(* Logix 5000 project; controller _GigaDiscovery vendor 1 type 14 code 244 rev 35.11; software revision 35.03; part 8 of 23 *)
(* tags used below, declared in another part *)
   ArmInductanceGondola : REAL;
   ArmResistanceGondola : REAL;
   First_Push_Angle : REAL;   // WEIGHT
   Gondola_Start_Delay : TIMER;
   Gondola_Stop : BOOL;
   Max_Torque_for_Angle_Correction : REAL;
   Min_error_to_Start_Decreasing_Torque : REAL;
   Os : DINT;
   Os_to_CCW : BOOL;
   Os_to_CW : BOOL;
   Pylon_Sequencer : Sequencer;
   SpeedRegKi : REAL;
   SpeedRegKp : REAL;
   Timer : TIMER[10];
   Angle_at_Full_Load : REAL;
   Angle_at_min_Load : REAL;
   AngleContrl : REAL;
   Auto_Cycle_Step : DINT;
   Braking_Torque_Lim : REAL;
   CurrentLimit : DINT;
   Direction : BOOL;   // 1 = Spinta CW 0 = Spinta CCW
   Enable_to_Start : UDT_CROUT;   // Abilitazione allo start QC8011E QC8013E
   Encoder_Resetted : BOOL;
   First_Push_Set_Torque_to_Zero : BOOL;
   Girella_Field_Actuate_During_Inactivity : BOOL;
   Gondola_Axe : Axe;
   Gondola_Decc_timer_Start : BOOL;
   Gondola_Immediatly_Stop : BOOL;
   Gondola_Out_Ref : INT;
   Gondola_Speed_Ref_ABS : REAL;
   Gondola_Speed_Reference : DINT;
   Gondola_Stop_CW : BOOL;   // Gondola Sto Direction 0 > CCW 1 > CW
   Gondola_Stop_Step : DINT;
   HMI_Gondola_Start_Delay : DINT;
   HMI_Overspeed_Test_Pb : BOOL;
   HMI_Reset_Encoder_Position : BOOL;
   I_Gondola_Home_Position_Sensor_1 : UDT_DCM;   // Home Sensor Speed Check -B40002I
   I_Pylon_Home_Ch1 : UDT_DCM;   // Home position Pylon Ch1 -B26002I
   I_Pylon_Home_Ch2 : UDT_DCM;   // Home position Pylon Ch2 -B26007I
   I_Zero_Set_Sensor : BOOL;   // Zero Set Sensor -B11201A
   Increase_Torque_Limit_Mem : BOOL;
   K_Brake : REAL;
   K_Speed_Factor : REAL;
   Max_Empty_Torque : REAL;   // 75
   Max_Full_Torque : REAL;   // 85
   MAX_HMI_Speed_Value : DINT;
   Max_Reference_Output : DINT;
   Max_Speed_Reference : DINT;
   Min_Speed_Reference : DINT;
   Min_Torque_to_Maintain_Height_Full_Load : REAL;
   Min_Torque_to_Maintain_Height_min_Load : REAL;
   No_Sfty : Std_to_Sfty;
   Os_to_CW_CCW : BOOL;
   Oscillation_Error : REAL;
   Pylon_Axe : Axe;
   Pylon_Field_Actuate_During_Inactivity : BOOL;
   Pylon_Filtered_Speed : REAL;
   Pylon_Reference : DINT;
   Ratio_HMI_Speed_Ref : REAL;
   Reference_Out_Conversion_Pylon : REAL;
   Reset_Pulse : BOOL;
   RPM_Max_Motor_Speed_Pylon : DINT;
   Start_Stop_Cycle : Sequencer;
   Stop_Request : BOOL;
   Timers : TIMER[32];
   To_Sfty : Std_to_Sfty;
   Torque_Cmd_from_Cycle : REAL;
   TorqueNeg_Angle_Control : REAL;
   TorquePos_Angle_Control : REAL;
   Work_Auto_Cycle : Auto_Cycle;
(* Pylon, continued *)

ROUTINE _02_Ctrl_Mode   (* ladder *)
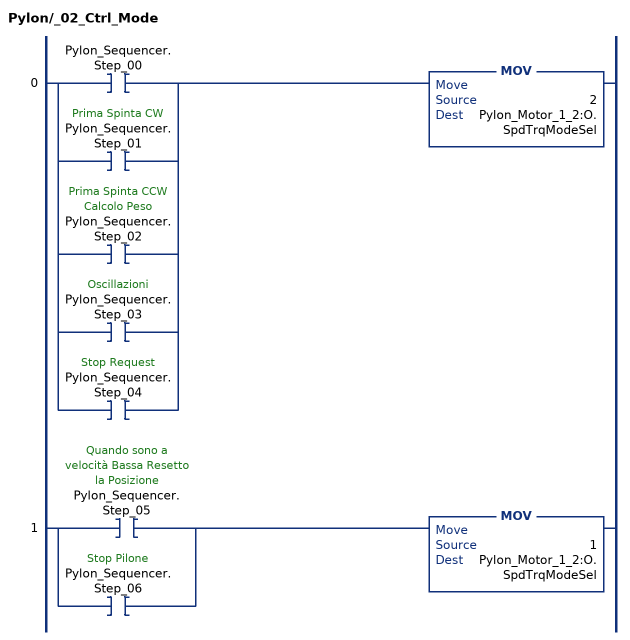
   0: [XIC(Pylon_Sequencer.Step_00) ,XIC(Pylon_Sequencer.Step_01) ,XIC(Pylon_Sequencer.Step_02) ,XIC(Pylon_Sequencer.Step_03) ,XIC(Pylon_Sequencer.Step_04) ]MOV(2,Pylon_Motor_1_2:O.SpdTrqModeSel);
   1: [XIC(Pylon_Sequencer.Step_05) ,XIC(Pylon_Sequencer.Step_06) ]MOV(1,Pylon_Motor_1_2:O.SpdTrqModeSel);
END_ROUTINE

ROUTINE _03_Speed_Ref   (* ladder *)
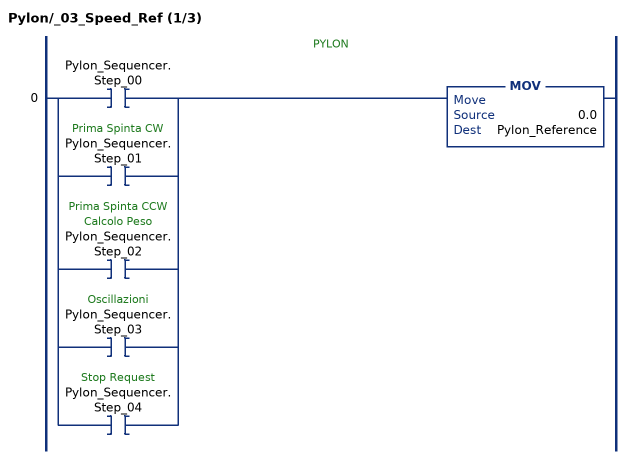
   // PYLON
   0: [XIC(Pylon_Sequencer.Step_00) ,XIC(Pylon_Sequencer.Step_01) ,XIC(Pylon_Sequencer.Step_02) ,XIC(Pylon_Sequencer.Step_03) ,XIC(Pylon_Sequencer.Step_04) ]MOV(0.0,Pylon_Reference);
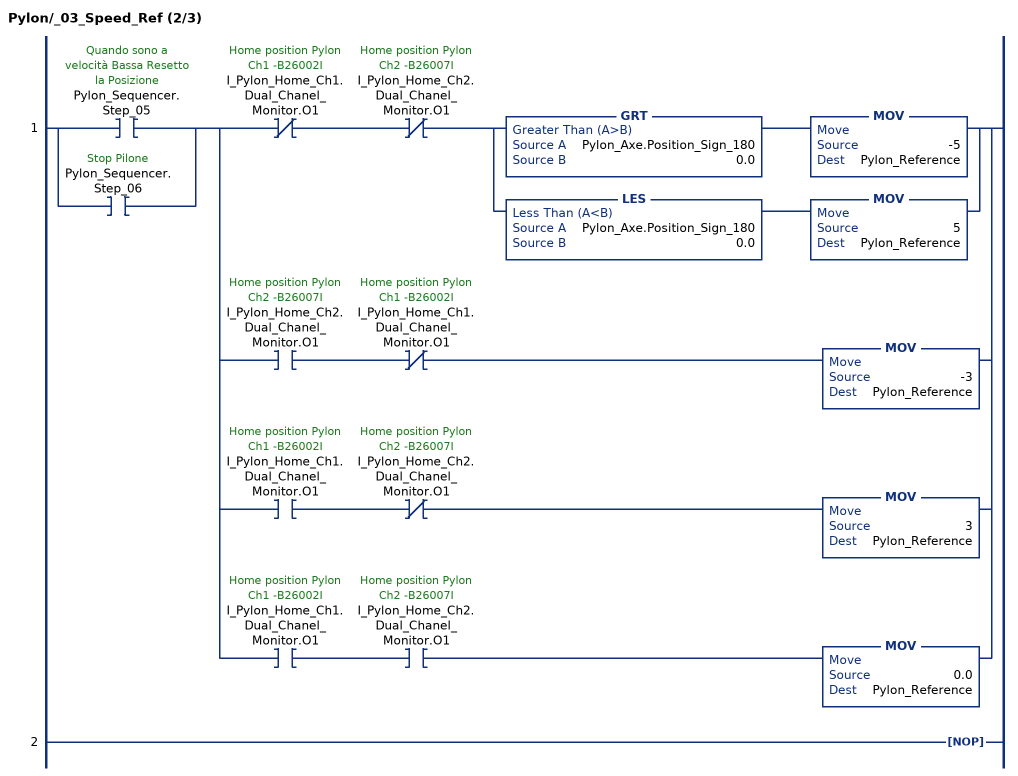
   1: [XIC(Pylon_Sequencer.Step_05) ,XIC(Pylon_Sequencer.Step_06) ][XIO(I_Pylon_Home_Ch1.Dual_Chanel_Monitor.O1) XIO(I_Pylon_Home_Ch2.Dual_Chanel_Monitor.O1) [GRT(Pylon_Axe.Position_Sign_180,0.0) MOV(-5,Pylon_Reference) ,LES(Pylon_Axe.Position_Sign_180,0.0) MOV(5,Pylon_Reference) ] ,[XIC(I_Pylon_Home_Ch2.Dual_Chanel_Monitor.O1) XIO(I_Pylon_Home_Ch1.Dual_Chanel_Monitor.O1) MOV(-3,Pylon_Reference) ,XIC(I_Pylon_Home_Ch1.Dual_Chanel_Monitor.O1) XIO(I_Pylon_Home_Ch2.Dual_Chanel_Monitor.O1) MOV(3,Pylon_Reference) ,XIC(I_Pylon_Home_Ch1.Dual_Chanel_Monitor.O1) XIC(I_Pylon_Home_Ch2.Dual_Chanel_Monitor.O1) MOV(0.0,Pylon_Reference) ] ];
   2: NOP();
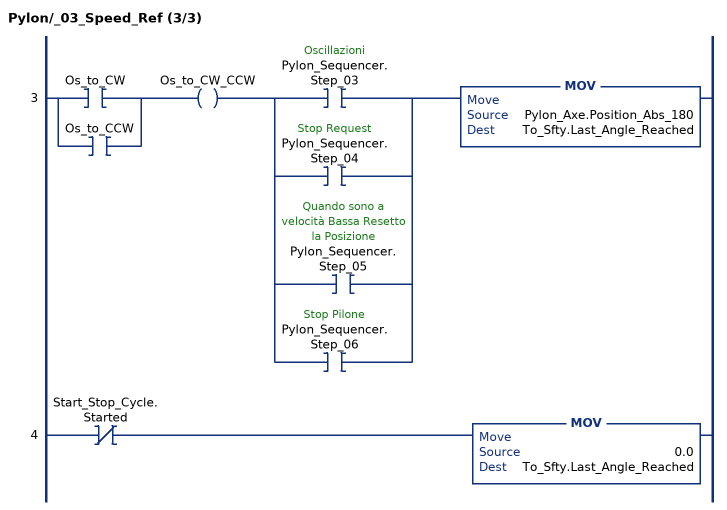
   3: [XIC(Os_to_CW) ,XIC(Os_to_CCW) ]OTE(Os_to_CW_CCW)[XIC(Pylon_Sequencer.Step_03) ,XIC(Pylon_Sequencer.Step_04) ,XIC(Pylon_Sequencer.Step_05) ,XIC(Pylon_Sequencer.Step_06) ]MOV(Pylon_Axe.Position_Abs_180,To_Sfty.Last_Angle_Reached);
   4: XIO(Start_Stop_Cycle.Started)MOV(0.0,To_Sfty.Last_Angle_Reached);
END_ROUTINE

ROUTINE _04_Torque_Lim   (* ladder *)
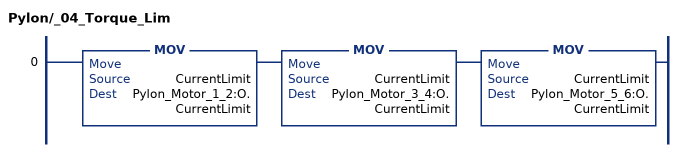
   0: MOV(CurrentLimit,Pylon_Motor_1_2:O.CurrentLimit)MOV(CurrentLimit,Pylon_Motor_3_4:O.CurrentLimit)MOV(CurrentLimit,Pylon_Motor_5_6:O.CurrentLimit);
END_ROUTINE

ROUTINE _05_Oscillation   (* ladder *)
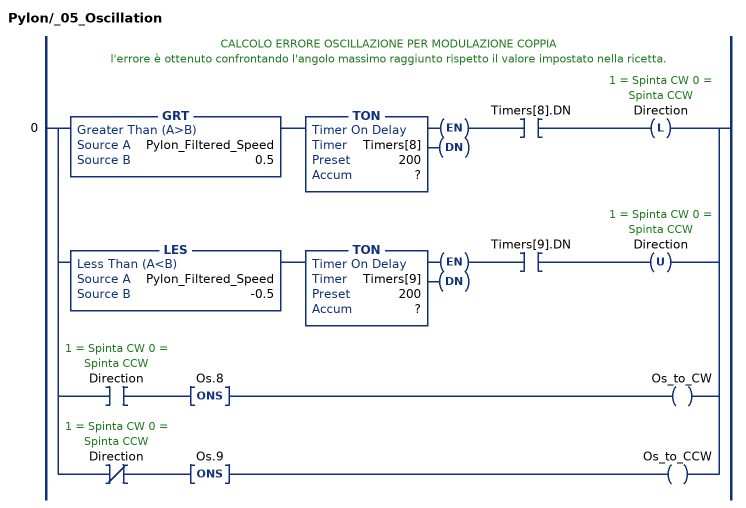
   // CALCOLO ERRORE OSCILLAZIONE PER MODULAZIONE COPPIA
   // l'errore è ottenuto confrontando l'angolo massimo raggiunto rispetto il valore impostato nella ricetta.
   0: [GRT(Pylon_Filtered_Speed,0.5) TON(Timers[8],?,?) XIC(Timers[8].DN) OTL(Direction) ,LES(Pylon_Filtered_Speed,-0.5) TON(Timers[9],?,?) XIC(Timers[9].DN) OTU(Direction) ,XIC(Direction) ONS(Os.8) OTE(Os_to_CW) ,XIO(Direction) ONS(Os.9) OTE(Os_to_CCW) ];
END_ROUTINE

ROUTINE _06_Scale_Angle   (* function block diagram *)
   SHEET 1
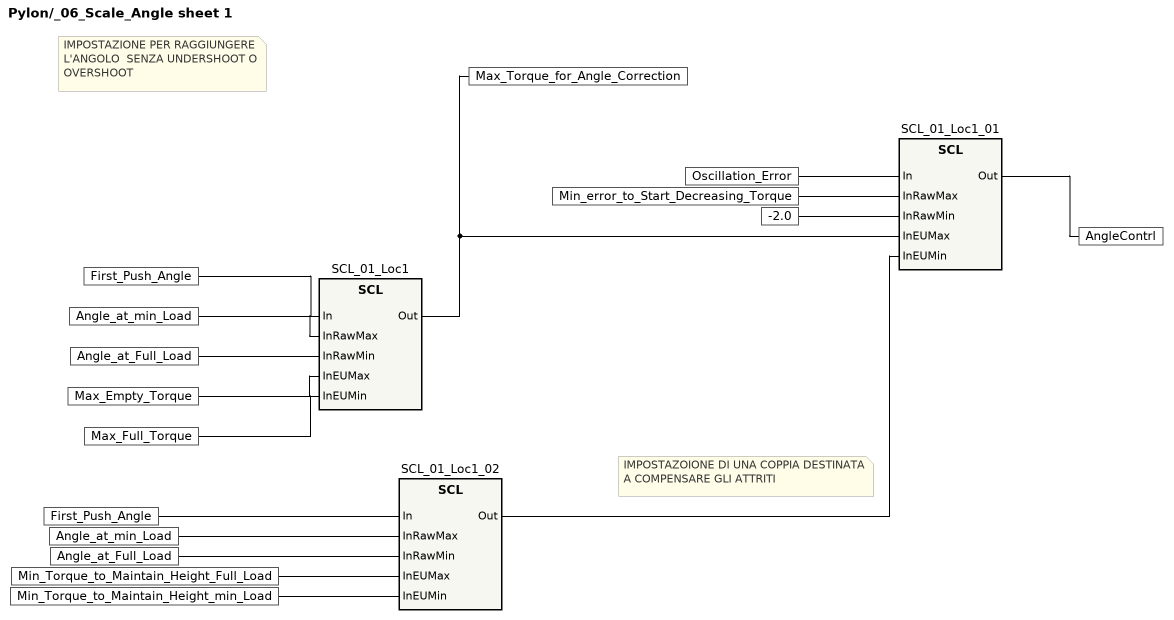
   // IMPOSTAZIONE PER RAGGIUNGERE
   // L'ANGOLO  SENZA UNDERSHOOT O
   // OVERSHOOT
   SCL_01_Loc1 : SCL(In := First_Push_Angle, InRawMax := Angle_at_min_Load, InRawMin := Angle_at_Full_Load, InEUMax := Max_Empty_Torque, InEUMin := Max_Full_Torque);
   // IMPOSTAZOIONE DI UNA COPPIA DESTINATA
   // A COMPENSARE GLI ATTRITI
   SCL_01_Loc1_02 : SCL(In := First_Push_Angle, InRawMax := Angle_at_min_Load, InRawMin := Angle_at_Full_Load, InEUMax := Min_Torque_to_Maintain_Height_Full_Load, InEUMin := Min_Torque_to_Maintain_Height_min_Load);
   Max_Torque_for_Angle_Correction := SCL_01_Loc1.Out;
   SCL_01_Loc1_01 : SCL(In := Oscillation_Error, InRawMax := Min_error_to_Start_Decreasing_Torque, InRawMin := -2.0, InEUMax := SCL_01_Loc1.Out, InEUMin := SCL_01_Loc1_02.Out);
   AngleContrl := SCL_01_Loc1_01.Out;
END_ROUTINE

ROUTINE _07_Torque_Cmd   (* ladder *)
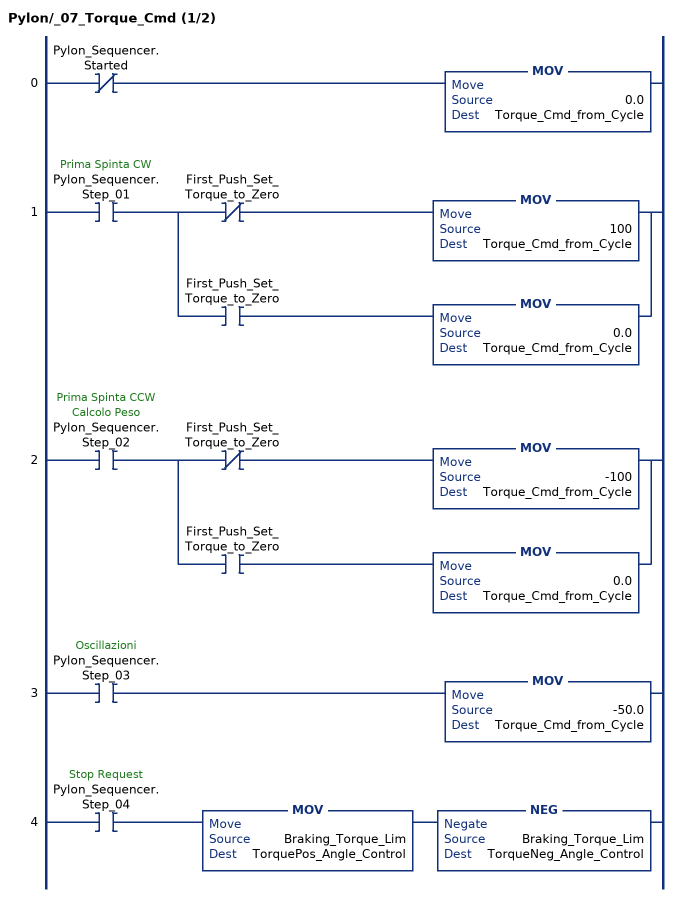
   0: XIO(Pylon_Sequencer.Started)MOV(0.0,Torque_Cmd_from_Cycle);
   1: XIC(Pylon_Sequencer.Step_01)[XIO(First_Push_Set_Torque_to_Zero) MOV(100,Torque_Cmd_from_Cycle) ,XIC(First_Push_Set_Torque_to_Zero) MOV(0.0,Torque_Cmd_from_Cycle) ];
   2: XIC(Pylon_Sequencer.Step_02)[XIO(First_Push_Set_Torque_to_Zero) MOV(-100,Torque_Cmd_from_Cycle) ,XIC(First_Push_Set_Torque_to_Zero) MOV(0.0,Torque_Cmd_from_Cycle) ];
   3: XIC(Pylon_Sequencer.Step_03)MOV(-50.0,Torque_Cmd_from_Cycle);
   4: XIC(Pylon_Sequencer.Step_04)MOV(Braking_Torque_Lim,TorquePos_Angle_Control)NEG(Braking_Torque_Lim,TorqueNeg_Angle_Control);
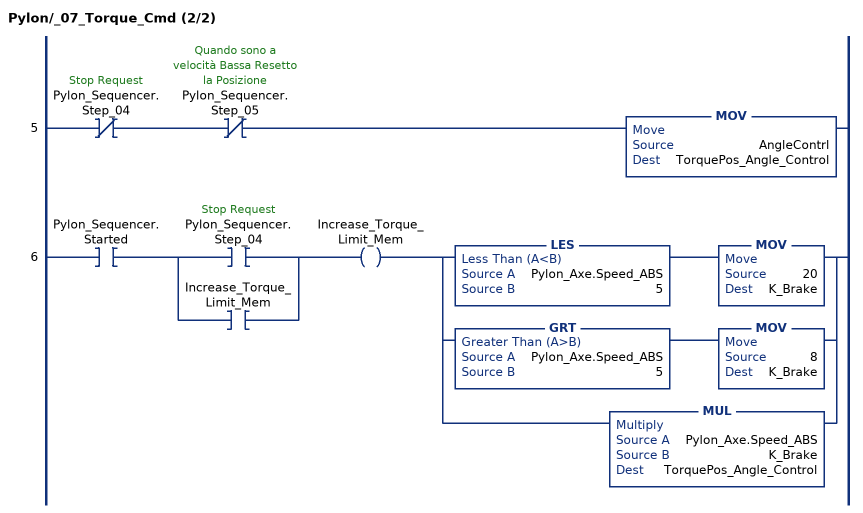
   5: XIO(Pylon_Sequencer.Step_04)XIO(Pylon_Sequencer.Step_05)MOV(AngleContrl,TorquePos_Angle_Control);
   6: XIC(Pylon_Sequencer.Started)[XIC(Pylon_Sequencer.Step_04) ,XIC(Increase_Torque_Limit_Mem) ]OTE(Increase_Torque_Limit_Mem)[LES(Pylon_Axe.Speed_ABS,5) MOV(20,K_Brake) ,GRT(Pylon_Axe.Speed_ABS,5) MOV(8,K_Brake) ,MUL(Pylon_Axe.Speed_ABS,K_Brake,TorquePos_Angle_Control) ];
END_ROUTINE

ROUTINE _08_Gondola   (* ladder *)
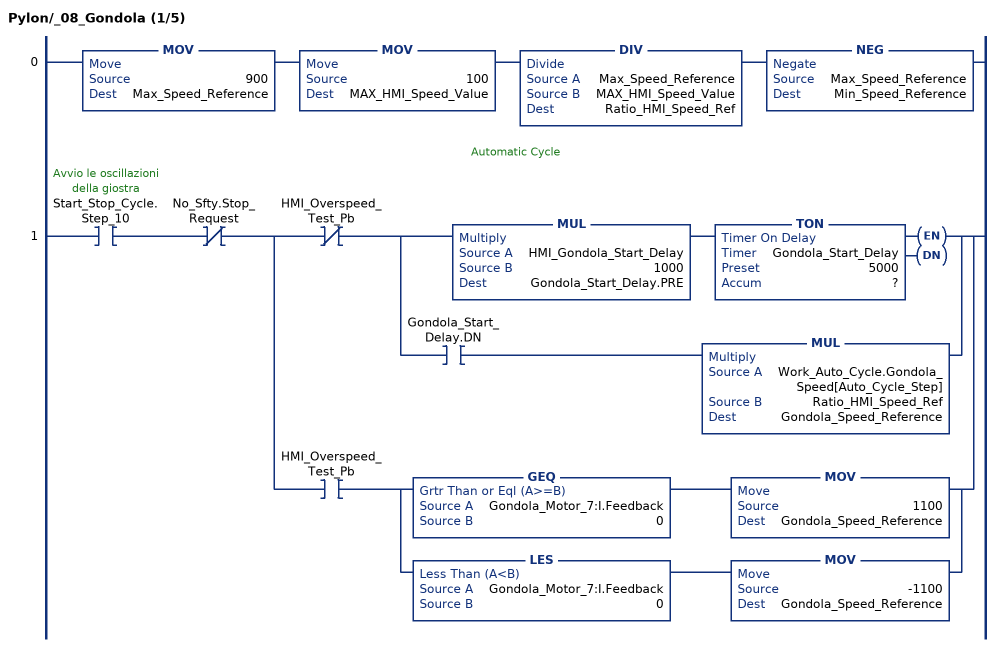
   0: MOV(900,Max_Speed_Reference)MOV(100,MAX_HMI_Speed_Value)DIV(Max_Speed_Reference,MAX_HMI_Speed_Value,Ratio_HMI_Speed_Ref)NEG(Max_Speed_Reference,Min_Speed_Reference);
   // Automatic Cycle
   1: XIC(Start_Stop_Cycle.Step_10)XIO(No_Sfty.Stop_Request)[XIO(HMI_Overspeed_Test_Pb) [MUL(HMI_Gondola_Start_Delay,1000,Gondola_Start_Delay.PRE) TON(Gondola_Start_Delay,?,?) ,XIC(Gondola_Start_Delay.DN) MUL(Work_Auto_Cycle.Gondola_Speed[Auto_Cycle_Step],Ratio_HMI_Speed_Ref,Gondola_Speed_Reference) ] ,XIC(HMI_Overspeed_Test_Pb) [GEQ(Gondola_Motor_7:I.Feedback,0) MOV(1100,Gondola_Speed_Reference) ,LES(Gondola_Motor_7:I.Feedback,0) MOV(-1100,Gondola_Speed_Reference) ] ];
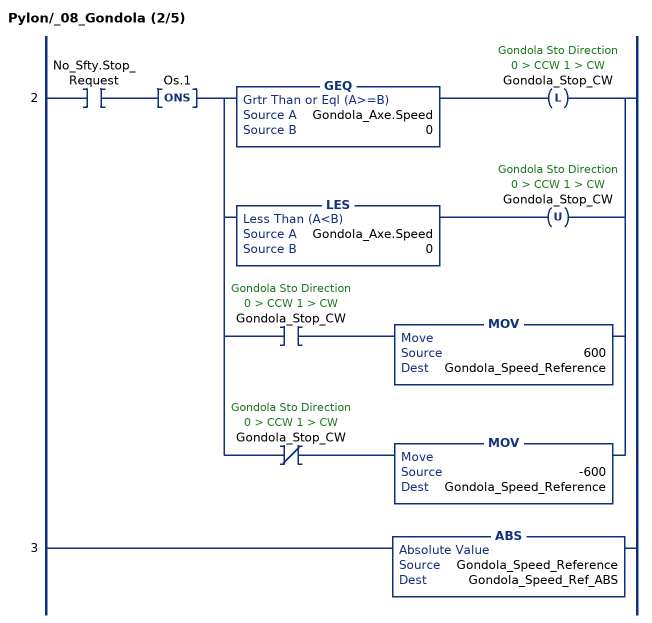
   2: XIC(No_Sfty.Stop_Request)ONS(Os.1)[GEQ(Gondola_Axe.Speed,0) OTL(Gondola_Stop_CW) ,LES(Gondola_Axe.Speed,0) OTU(Gondola_Stop_CW) ,XIC(Gondola_Stop_CW) MOV(600,Gondola_Speed_Reference) ,XIO(Gondola_Stop_CW) MOV(-600,Gondola_Speed_Reference) ];
   3: ABS(Gondola_Speed_Reference,Gondola_Speed_Ref_ABS);
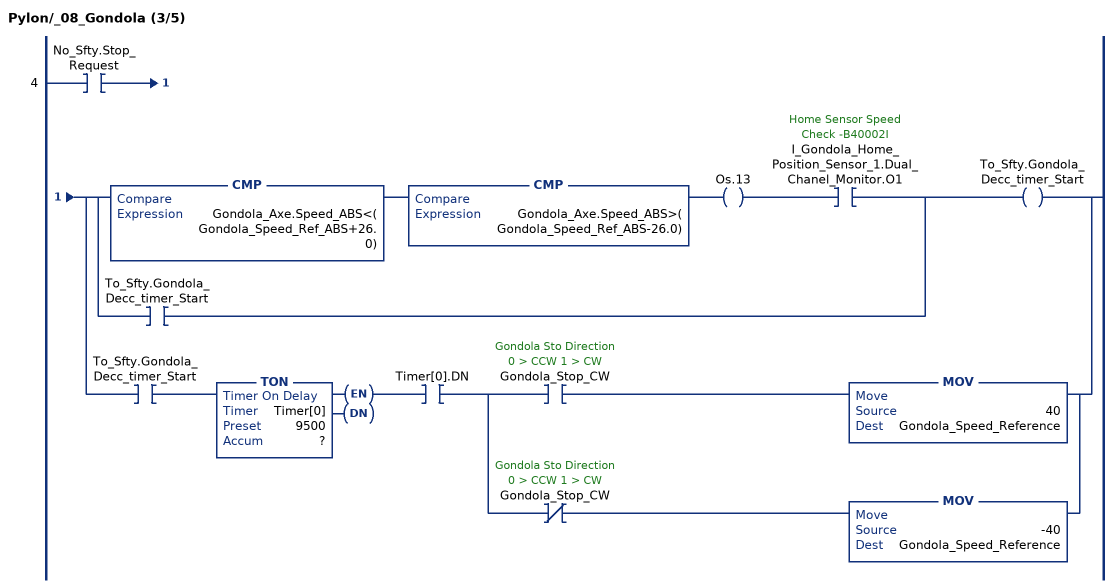
   4: XIC(No_Sfty.Stop_Request)[[CMP(Gondola_Axe.Speed_ABS<(Gondola_Speed_Ref_ABS+26.0)) CMP(Gondola_Axe.Speed_ABS>(Gondola_Speed_Ref_ABS-26.0)) OTE(Os.13) XIC(I_Gondola_Home_Position_Sensor_1.Dual_Chanel_Monitor.O1) ,XIC(To_Sfty.Gondola_Decc_timer_Start) ] OTE(To_Sfty.Gondola_Decc_timer_Start) ,XIC(To_Sfty.Gondola_Decc_timer_Start) TON(Timer[0],?,?) XIC(Timer[0].DN) [XIC(Gondola_Stop_CW) MOV(40,Gondola_Speed_Reference) ,XIO(Gondola_Stop_CW) MOV(-40,Gondola_Speed_Reference) ] ];
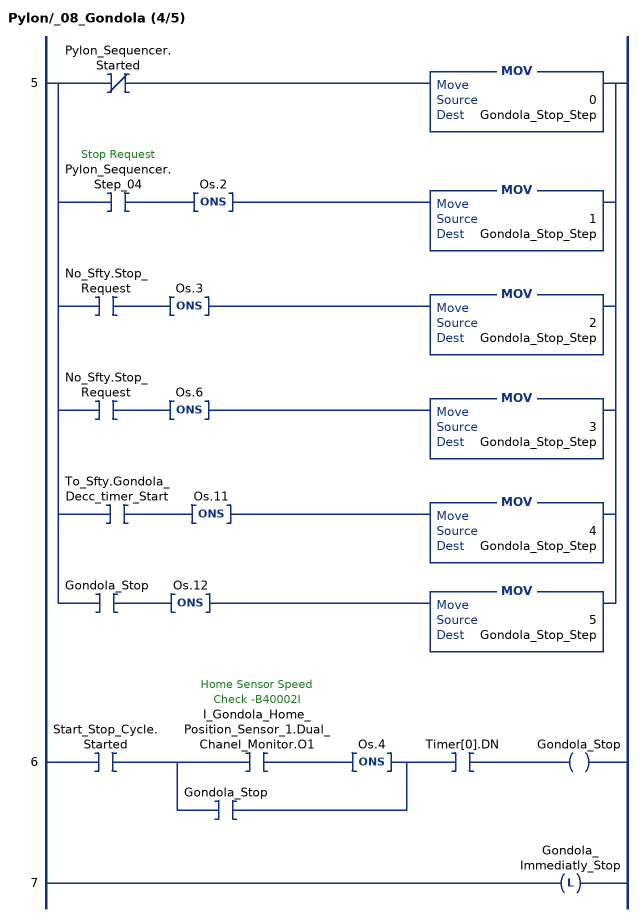
   5: [XIO(Pylon_Sequencer.Started) MOV(0,Gondola_Stop_Step) ,XIC(Pylon_Sequencer.Step_04) ONS(Os.2) MOV(1,Gondola_Stop_Step) ,XIC(No_Sfty.Stop_Request) ONS(Os.3) MOV(2,Gondola_Stop_Step) ,XIC(No_Sfty.Stop_Request) ONS(Os.6) MOV(3,Gondola_Stop_Step) ,XIC(To_Sfty.Gondola_Decc_timer_Start) ONS(Os.11) MOV(4,Gondola_Stop_Step) ,XIC(Gondola_Stop) ONS(Os.12) MOV(5,Gondola_Stop_Step) ];
   6: XIC(Start_Stop_Cycle.Started)[XIC(I_Gondola_Home_Position_Sensor_1.Dual_Chanel_Monitor.O1) ONS(Os.4) ,XIC(Gondola_Stop) ]XIC(Timer[0].DN)OTE(Gondola_Stop);
   7: OTL(Gondola_Immediatly_Stop);
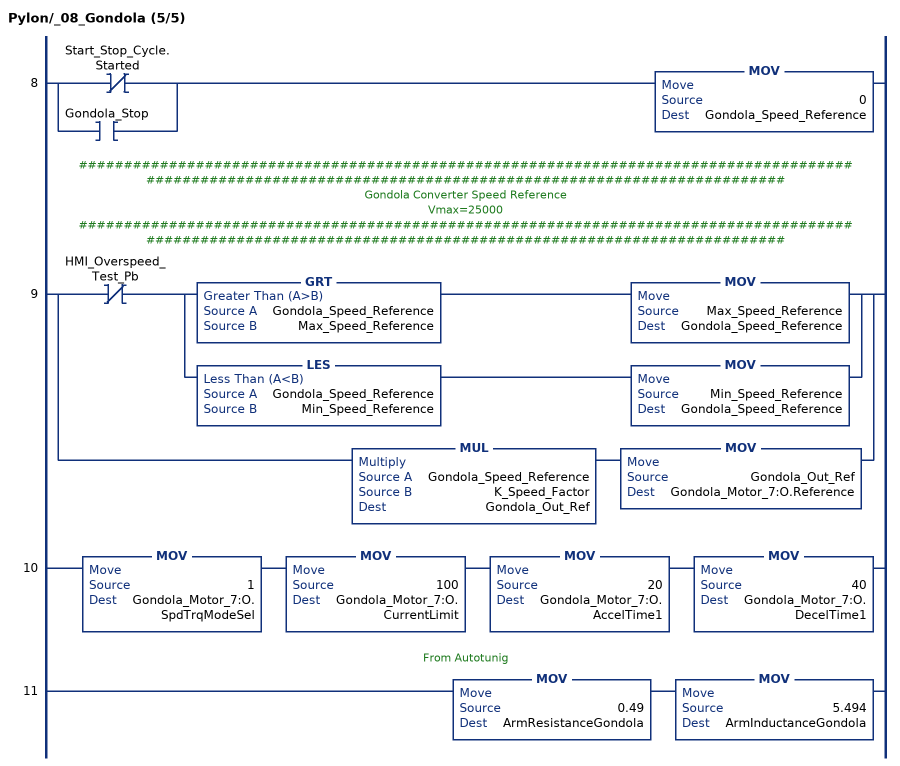
   8: [XIO(Start_Stop_Cycle.Started) ,XIC(Gondola_Stop) ]MOV(0,Gondola_Speed_Reference);
   // #############################################################################################################################################################
   // Gondola Converter Speed Reference
   // Vmax=25000
   // #############################################################################################################################################################
   9: [XIO(HMI_Overspeed_Test_Pb) [GRT(Gondola_Speed_Reference,Max_Speed_Reference) MOV(Max_Speed_Reference,Gondola_Speed_Reference) ,LES(Gondola_Speed_Reference,Min_Speed_Reference) MOV(Min_Speed_Reference,Gondola_Speed_Reference) ] ,MUL(Gondola_Speed_Reference,K_Speed_Factor,Gondola_Out_Ref) MOV(Gondola_Out_Ref,Gondola_Motor_7:O.Reference) ];
   10: MOV(1,Gondola_Motor_7:O.SpdTrqModeSel)MOV(100,Gondola_Motor_7:O.CurrentLimit)MOV(20,Gondola_Motor_7:O.AccelTime1)MOV(40,Gondola_Motor_7:O.DecelTime1);
   // From Autotunig
   11: MOV(0.49,ArmResistanceGondola)MOV(5.494,ArmInductanceGondola);
END_ROUTINE

ROUTINE _99_Drive_Commands   (* ladder *)
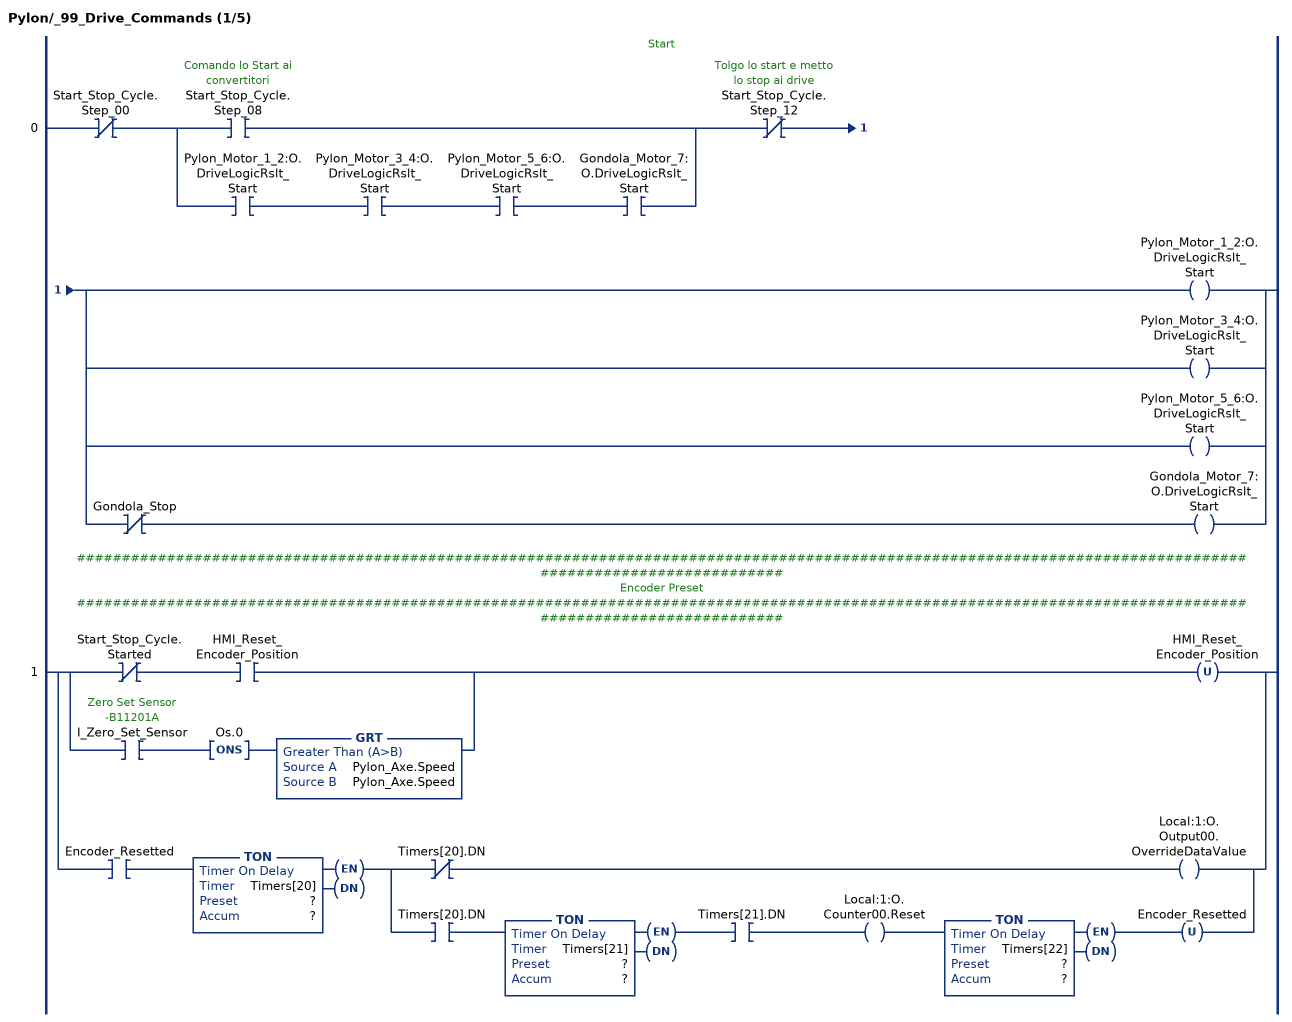
   // Start
   0: XIO(Start_Stop_Cycle.Step_00)[XIC(Start_Stop_Cycle.Step_08) ,XIC(Pylon_Motor_1_2:O.DriveLogicRslt_Start) XIC(Pylon_Motor_3_4:O.DriveLogicRslt_Start) XIC(Pylon_Motor_5_6:O.DriveLogicRslt_Start) XIC(Gondola_Motor_7:O.DriveLogicRslt_Start) ]XIO(Start_Stop_Cycle.Step_12)[OTE(Pylon_Motor_1_2:O.DriveLogicRslt_Start) ,OTE(Pylon_Motor_3_4:O.DriveLogicRslt_Start) ,OTE(Pylon_Motor_5_6:O.DriveLogicRslt_Start) ,XIO(Gondola_Stop) OTE(Gondola_Motor_7:O.DriveLogicRslt_Start) ];
   // #############################################################################################################################################################
   // Encoder Preset
   // #############################################################################################################################################################
   1: [[XIO(Start_Stop_Cycle.Started) XIC(HMI_Reset_Encoder_Position) ,XIC(I_Zero_Set_Sensor) ONS(Os.0) GRT(Pylon_Axe.Speed,Pylon_Axe.Speed) ] OTU(HMI_Reset_Encoder_Position) ,XIC(Encoder_Resetted) TON(Timers[20],?,?) [XIO(Timers[20].DN) OTE(Local:1:O.Output00.OverrideDataValue) ,XIC(Timers[20].DN) TON(Timers[21],?,?) XIC(Timers[21].DN) OTE(Local:1:O.Counter00.Reset) TON(Timers[22],?,?) OTU(Encoder_Resetted) ] ];
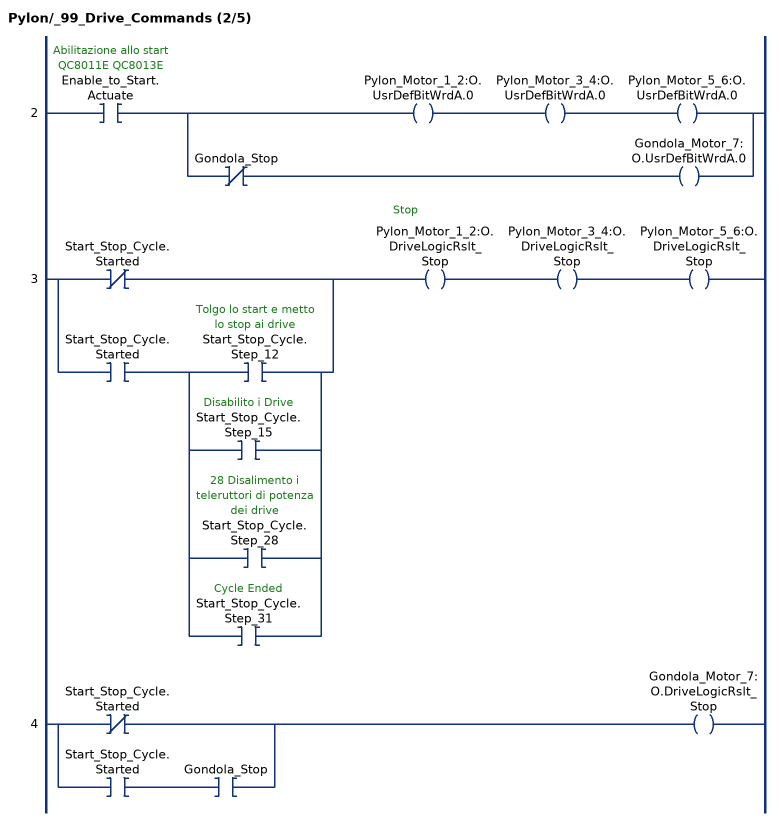
   2: XIC(Enable_to_Start.Actuate)[OTE(Pylon_Motor_1_2:O.UsrDefBitWrdA.0) OTE(Pylon_Motor_3_4:O.UsrDefBitWrdA.0) OTE(Pylon_Motor_5_6:O.UsrDefBitWrdA.0) ,XIO(Gondola_Stop) OTE(Gondola_Motor_7:O.UsrDefBitWrdA.0) ];
   // Stop
   3: [XIO(Start_Stop_Cycle.Started) ,XIC(Start_Stop_Cycle.Started) [XIC(Start_Stop_Cycle.Step_12) ,XIC(Start_Stop_Cycle.Step_15) ,XIC(Start_Stop_Cycle.Step_28) ,XIC(Start_Stop_Cycle.Step_31) ] ]OTE(Pylon_Motor_1_2:O.DriveLogicRslt_Stop)OTE(Pylon_Motor_3_4:O.DriveLogicRslt_Stop)OTE(Pylon_Motor_5_6:O.DriveLogicRslt_Stop);
   4: [XIO(Start_Stop_Cycle.Started) ,XIC(Start_Stop_Cycle.Started) XIC(Gondola_Stop) ]OTE(Gondola_Motor_7:O.DriveLogicRslt_Stop);
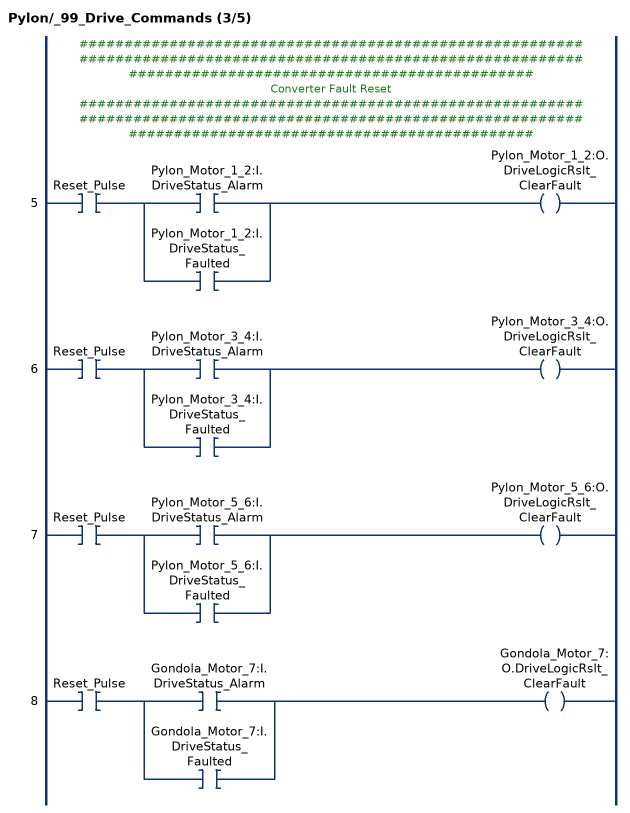
   // #############################################################################################################################################################
   // Converter Fault Reset
   // #############################################################################################################################################################
   5: XIC(Reset_Pulse)[XIC(Pylon_Motor_1_2:I.DriveStatus_Alarm) ,XIC(Pylon_Motor_1_2:I.DriveStatus_Faulted) ]OTE(Pylon_Motor_1_2:O.DriveLogicRslt_ClearFault);
   6: XIC(Reset_Pulse)[XIC(Pylon_Motor_3_4:I.DriveStatus_Alarm) ,XIC(Pylon_Motor_3_4:I.DriveStatus_Faulted) ]OTE(Pylon_Motor_3_4:O.DriveLogicRslt_ClearFault);
   7: XIC(Reset_Pulse)[XIC(Pylon_Motor_5_6:I.DriveStatus_Alarm) ,XIC(Pylon_Motor_5_6:I.DriveStatus_Faulted) ]OTE(Pylon_Motor_5_6:O.DriveLogicRslt_ClearFault);
   8: XIC(Reset_Pulse)[XIC(Gondola_Motor_7:I.DriveStatus_Alarm) ,XIC(Gondola_Motor_7:I.DriveStatus_Faulted) ]OTE(Gondola_Motor_7:O.DriveLogicRslt_ClearFault);
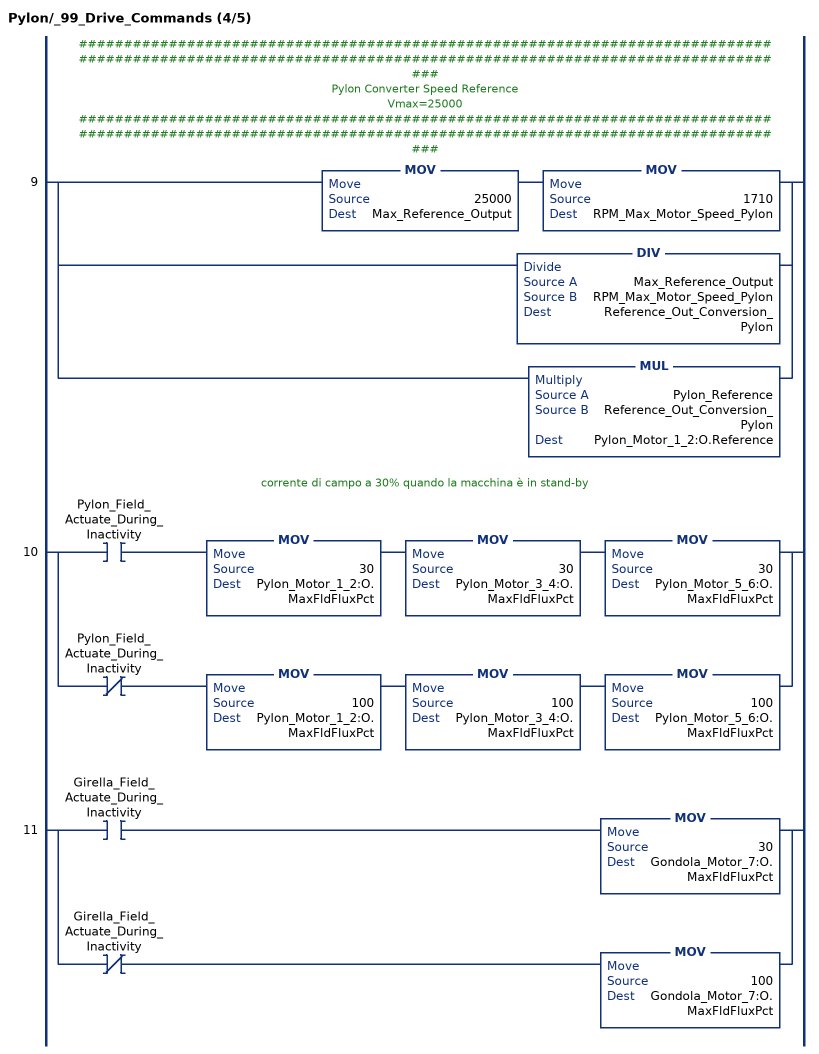
   // #############################################################################################################################################################
   // Pylon Converter Speed Reference
   // Vmax=25000
   // #############################################################################################################################################################
   9: [MOV(25000,Max_Reference_Output) MOV(1710,RPM_Max_Motor_Speed_Pylon) ,DIV(Max_Reference_Output,RPM_Max_Motor_Speed_Pylon,Reference_Out_Conversion_Pylon) ,MUL(Pylon_Reference,Reference_Out_Conversion_Pylon,Pylon_Motor_1_2:O.Reference) ];
   // corrente di campo a 30% quando la macchina è in stand-by
   10: [XIC(Pylon_Field_Actuate_During_Inactivity) MOV(30,Pylon_Motor_1_2:O.MaxFldFluxPct) MOV(30,Pylon_Motor_3_4:O.MaxFldFluxPct) MOV(30,Pylon_Motor_5_6:O.MaxFldFluxPct) ,XIO(Pylon_Field_Actuate_During_Inactivity) MOV(100,Pylon_Motor_1_2:O.MaxFldFluxPct) MOV(100,Pylon_Motor_3_4:O.MaxFldFluxPct) MOV(100,Pylon_Motor_5_6:O.MaxFldFluxPct) ];
   11: [XIC(Girella_Field_Actuate_During_Inactivity) MOV(30,Gondola_Motor_7:O.MaxFldFluxPct) ,XIO(Girella_Field_Actuate_During_Inactivity) MOV(100,Gondola_Motor_7:O.MaxFldFluxPct) ];
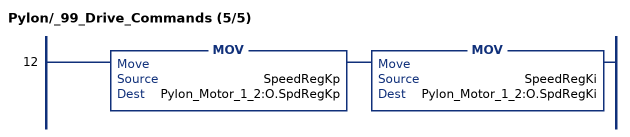
   12: MOV(SpeedRegKp,Pylon_Motor_1_2:O.SpdRegKp)MOV(SpeedRegKi,Pylon_Motor_1_2:O.SpdRegKi);
END_ROUTINE
